screen "St_Time machine data_4" 320x240
   IOField "I/O field_13" at 243,83 size 56x19; FormatPattern 999.99; Unit   %
      ProcessValue <- "Data_Real_%Mesin Stop[4]"
   IOField "I/O field_14" at 243,101 size 56x19; FormatPattern 999.99; Unit   %
      ProcessValue <- "Data_Real_%Mesin Run Baypass[4]"
   IOField "I/O field_11" at 243,66 size 56x19; FormatPattern 999.99; Unit   %
      ProcessValue <- "Data_Real_%Mesin Run[4]"
   Button "Button_1" at 46,213 size 90x25; TextOff 'Statistic Data'
      on Click: ActivateScreen("St_Data Statistic", 0)
   Button "Button_3" at 1,213 size 41x25; TextOff 'Main Page'; PictureOff "Home"
      on Click: ActivateScreen("Main Page", 0)
   Button "Button_2" at 237,213 size 80x25; TextOff 'Next page -->'; TextOn 'Page 3'
      on Click: ActivateScreen("St_Error Counter_4", 0)
   TextField "Text field_1" at 3,0 size 155x18; Text 'CURRENT SHIFT MINUS 4'
   TextField "Text field_31" at 7,101 size 21x19; Text '3'
   TextField "Text field_30" at 7,83 size 21x19; Text '2'
   TextField "Text field_29" at 7,66 size 21x19; Text '1'
   TextField "Text field_28" at 7,48 size 21x19; Text 'No'
   IOField "I/O field_21" at 219,83 size 25x19; FormatPattern 999
      ProcessValue <- "Data_DTLData_DTL_Mesin Stop[4].SECOND"
   IOField "I/O field_22" at 195,83 size 25x19; FormatPattern 999
      ProcessValue <- "Data_DTLData_DTL_Mesin Stop[4].MINUTE"
   IOField "I/O field_23" at 171,84 size 25x19; FormatPattern 999
      ProcessValue <- "Data_DTLData_DTL_Mesin Stop[4].HOUR"
   TextField "Text field_25" at 27,83 size 145x19; Text 'Stop'
   IOField "I/O field_4" at 219,101 size 25x19; FormatPattern 999
      ProcessValue <- "Data_DTLData_DTL_Mesin Run Baypass[4].SECOND"
   IOField "I/O field_5" at 195,101 size 25x19; FormatPattern 999
      ProcessValue <- "Data_DTLData_DTL_Mesin Run Baypass[4].MINUTE"
   IOField "I/O field_9" at 171,101 size 25x19; FormatPattern 999
      ProcessValue <- "Data_DTLData_DTL_Mesin Run Baypass[4].HOUR"
   TextField "Text field_12" at 219,48 size 25x19; Text 'Sec'
   TextField "Text field_11" at 195,48 size 25x19; Text 'Min'
   IOField "I/O field_2" at 219,66 size 25x19; FormatPattern 999
      ProcessValue <- "Data_DTLData_DTL_Mesin Run[4].SECOND"
   IOField "I/O field_3" at 195,66 size 25x19; FormatPattern 999
      ProcessValue <- "Data_DTLData_DTL_Mesin Run[4].MINUTE"
   TextField "Text field_3" at 27,48 size 145x19; Text 'Time Counter Machine'
   TextField "Text field_4" at 27,66 size 145x19; Text 'Running'
   TextField "Text field_5" at 27,101 size 145x19; Text 'Running Bypass'
   IOField "I/O field_24" at 171,66 size 25x19; FormatPattern 999
      ProcessValue <- "Data_DTLData_DTL_Mesin Run[4].HOUR"
   Button "Button_4" at 151,213 size 80x25; TextOff '<-- Back Page'; TextOn 'Page 1'
      on Click: ActivateScreen("St_Quantity Data_4", 0)
   TextField "Text field_6" at 260,0 size 57x15; Text 'Page 2 of 3'
   IOField "I/O field_1" at 243,119 size 56x19; FormatPattern 999.99; Unit   %
      ProcessValue <- "Data_Real_%Mesin Error[4]"
   TextField "Text field_7" at 7,119 size 21x19; Text '4'
   IOField "I/O field_8" at 219,119 size 25x19; FormatPattern 999
      ProcessValue <- "Data_DTLData_DTL_Mesin Error[4].SECOND"
   IOField "I/O field_10" at 195,119 size 25x19; FormatPattern 999
      ProcessValue <- "Data_DTLData_DTL_Mesin Error[4].MINUTE"
   IOField "I/O field_12" at 171,119 size 25x19; FormatPattern 999
      ProcessValue <- "Data_DTLData_DTL_Mesin Error[4].HOUR"
   TextField "Text field_8" at 27,119 size 145x19; Text 'Error'
   TextField "Text field_2" at 171,48 size 25x19; Text 'Hour'
   IOField "I/O field_6" at 6,17 size 109x15; FormatPattern 9999999999999999999999999999999999999999
      ProcessValue <- "Data_DTL1_Cur_ShiftA_4"
   TextField "Text field_9" at 120,17 size 18x13; Text 'S/D'
   IOField "I/O field_7" at 143,17 size 109x15; FormatPattern 9999999999999999999999999999999999999999
      ProcessValue <- "Data_DTL1_Cur_ShiftB_4"
   IOField "I/O field_16" at 219,138 size 25x19; FormatPattern 999
      ProcessValue <- "Data_DTLData_Total Time Machine[4].SECOND"
   IOField "I/O field_17" at 195,138 size 25x19; FormatPattern 999
      ProcessValue <- "Data_DTLData_Total Time Machine[4].MINUTE"
   IOField "I/O field_18" at 171,138 size 25x19; FormatPattern 999
      ProcessValue <- "Data_DTLData_Total Time Machine[4].HOUR"
   TextField "Text field_10" at 27,138 size 145x19; Text 'Total'
   IOField "I/O field_27" at 253,16 size 66x17; FormatPattern ????????
      ProcessValue <- "Data_String_sDT_Machine id"

screen "St_Time machine data_5" 320x240
   IOField "I/O field_13" at 243,83 size 56x19; FormatPattern 999.99; Unit   %
      ProcessValue <- "Data_Real_%Mesin Stop[5]"
   IOField "I/O field_14" at 243,101 size 56x19; FormatPattern 999.99; Unit   %
      ProcessValue <- "Data_Real_%Mesin Run Baypass[5]"
   IOField "I/O field_11" at 243,66 size 56x19; FormatPattern 999.99; Unit   %
      ProcessValue <- "Data_Real_%Mesin Run[5]"
   Button "Button_1" at 46,213 size 90x25; TextOff 'Statistic Data'
      on Click: ActivateScreen("St_Data Statistic", 0)
   Button "Button_3" at 1,213 size 41x25; TextOff 'Main Page'; PictureOff "Home"
      on Click: ActivateScreen("Main Page", 0)
   Button "Button_2" at 237,213 size 80x25; TextOff 'Next page -->'; TextOn 'Page 3'
      on Click: ActivateScreen("St_Error Counter_5", 0)
   TextField "Text field_1" at 3,0 size 155x18; Text 'CURRENT SHIFT MINUS 5'
   TextField "Text field_31" at 7,101 size 21x19; Text '3'
   TextField "Text field_30" at 7,83 size 21x19; Text '2'
   TextField "Text field_29" at 7,66 size 21x19; Text '1'
   TextField "Text field_28" at 7,48 size 21x19; Text 'No'
   IOField "I/O field_21" at 219,83 size 25x19; FormatPattern 999
      ProcessValue <- "Data_DTLData_DTL_Mesin Stop[5].SECOND"
   IOField "I/O field_22" at 195,83 size 25x19; FormatPattern 999
      ProcessValue <- "Data_DTLData_DTL_Mesin Stop[5].MINUTE"
   IOField "I/O field_23" at 171,84 size 25x19; FormatPattern 999
      ProcessValue <- "Data_DTLData_DTL_Mesin Stop[5].HOUR"
   TextField "Text field_25" at 27,83 size 145x19; Text 'Stop'
   IOField "I/O field_4" at 219,101 size 25x19; FormatPattern 999
      ProcessValue <- "Data_DTLData_DTL_Mesin Run Baypass[5].SECOND"
   IOField "I/O field_5" at 195,101 size 25x19; FormatPattern 999
      ProcessValue <- "Data_DTLData_DTL_Mesin Run Baypass[5].MINUTE"
   IOField "I/O field_9" at 171,101 size 25x19; FormatPattern 999
      ProcessValue <- "Data_DTLData_DTL_Mesin Run Baypass[5].HOUR"
   TextField "Text field_12" at 219,48 size 25x19; Text 'Sec'
   TextField "Text field_11" at 195,48 size 25x19; Text 'Min'
   IOField "I/O field_2" at 219,66 size 25x19; FormatPattern 999
      ProcessValue <- "Data_DTLData_DTL_Mesin Run[5].SECOND"
   IOField "I/O field_3" at 195,66 size 25x19; FormatPattern 999
      ProcessValue <- "Data_DTLData_DTL_Mesin Run[5].MINUTE"
   TextField "Text field_3" at 27,48 size 145x19; Text 'Time Counter Machine'
   TextField "Text field_4" at 27,66 size 145x19; Text 'Running'
   TextField "Text field_5" at 27,101 size 145x19; Text 'Running Bypass'
   IOField "I/O field_24" at 171,66 size 25x19; FormatPattern 999
      ProcessValue <- "Data_DTLData_DTL_Mesin Run[5].HOUR"
   Button "Button_4" at 151,213 size 80x25; TextOff '<-- Back Page'; TextOn 'Page 1'
      on Click: ActivateScreen("St_Quantity Data_5", 0)
   TextField "Text field_6" at 260,0 size 57x15; Text 'Page 2 of 3'
   IOField "I/O field_1" at 243,119 size 56x19; FormatPattern 999.99; Unit   %
      ProcessValue <- "Data_Real_%Mesin Error[5]"
   TextField "Text field_7" at 7,119 size 21x19; Text '4'
   IOField "I/O field_8" at 219,119 size 25x19; FormatPattern 999
      ProcessValue <- "Data_DTLData_DTL_Mesin Error[5].SECOND"
   IOField "I/O field_10" at 195,119 size 25x19; FormatPattern 999
      ProcessValue <- "Data_DTLData_DTL_Mesin Error[5].MINUTE"
   IOField "I/O field_12" at 171,119 size 25x19; FormatPattern 999
      ProcessValue <- "Data_DTLData_DTL_Mesin Error[5].HOUR"
   TextField "Text field_8" at 27,119 size 145x19; Text 'Error'
   TextField "Text field_2" at 171,48 size 25x19; Text 'Hour'
   IOField "I/O field_6" at 6,17 size 109x15; FormatPattern 9999999999999999999999999999999999999999
      ProcessValue <- "Data_DTL1_Cur_ShiftA_5"
   TextField "Text field_9" at 120,17 size 18x13; Text 'S/D'
   IOField "I/O field_7" at 143,17 size 109x15; FormatPattern 9999999999999999999999999999999999999999
      ProcessValue <- "Data_DTL1_Cur_ShiftB_5"
   IOField "I/O field_16" at 219,138 size 25x19; FormatPattern 999
      ProcessValue <- "Data_DTLData_Total Time Machine[5].SECOND"
   IOField "I/O field_17" at 195,138 size 25x19; FormatPattern 999
      ProcessValue <- "Data_DTLData_Total Time Machine[5].MINUTE"
   IOField "I/O field_18" at 171,138 size 25x19; FormatPattern 999
      ProcessValue <- "Data_DTLData_Total Time Machine[5].HOUR"
   TextField "Text field_10" at 27,138 size 145x19; Text 'Total'
   IOField "I/O field_27" at 253,16 size 66x17; FormatPattern ????????
      ProcessValue <- "Data_String_sDT_Machine id"
*)